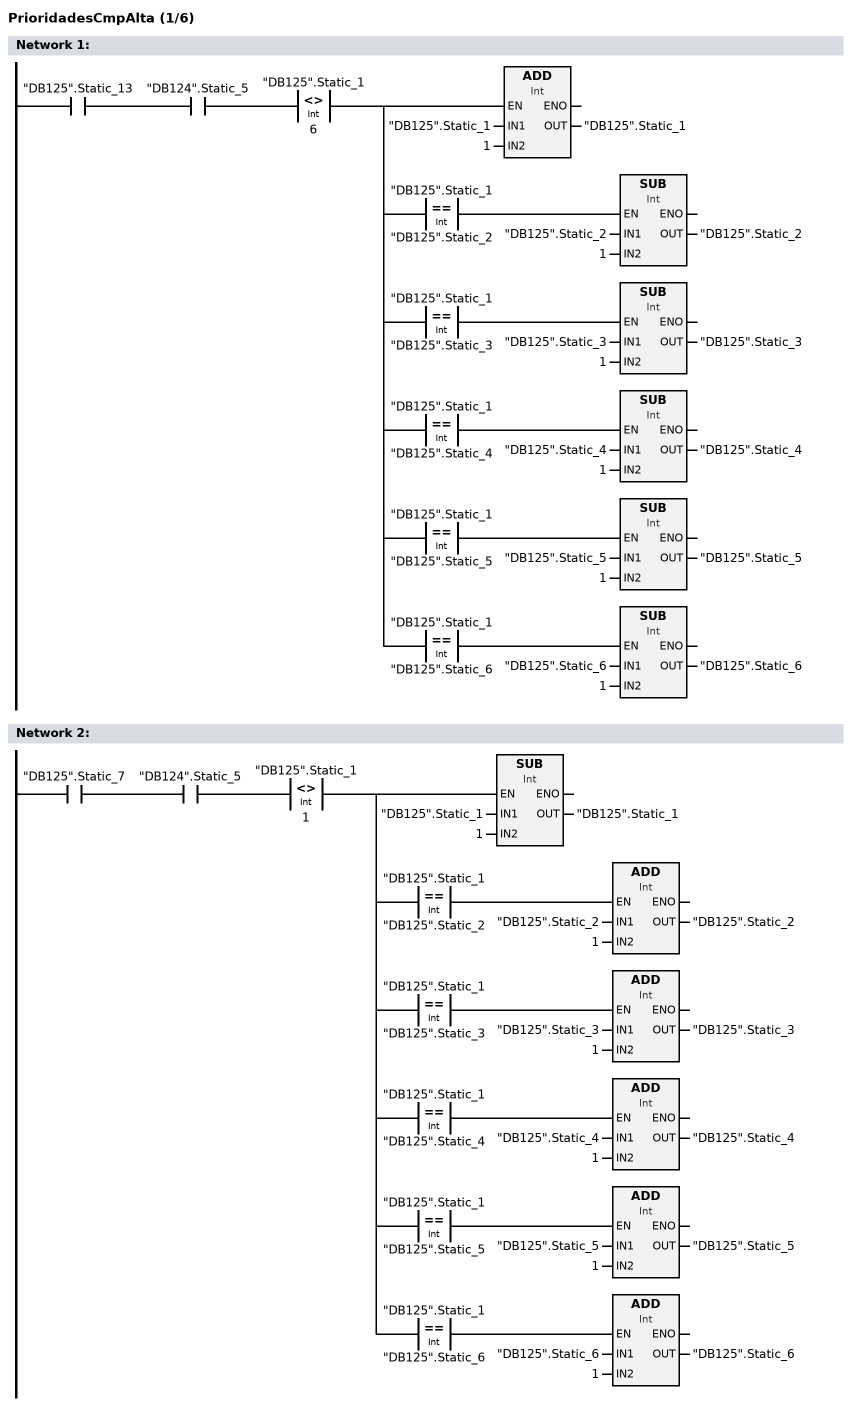
   #_w1 := "DB125".Static_13 AND "DB124".Static_5 AND ("DB125".Static_1 <> 6);
   IF #_w1 THEN "DB125".Static_1 := "DB125".Static_1 + 1; END_IF;
   IF #_w1 AND ("DB125".Static_1 = "DB125".Static_2) THEN "DB125".Static_2 := "DB125".Static_2 - 1; END_IF;
   IF #_w1 AND ("DB125".Static_1 = "DB125".Static_3) THEN "DB125".Static_3 := "DB125".Static_3 - 1; END_IF;
   IF #_w1 AND ("DB125".Static_1 = "DB125".Static_4) THEN "DB125".Static_4 := "DB125".Static_4 - 1; END_IF;
   IF #_w1 AND ("DB125".Static_1 = "DB125".Static_5) THEN "DB125".Static_5 := "DB125".Static_5 - 1; END_IF;
   IF #_w1 AND ("DB125".Static_1 = "DB125".Static_6) THEN "DB125".Static_6 := "DB125".Static_6 - 1; END_IF;
END_REGION

REGION Network 2
   #_w1 := "DB125".Static_7 AND "DB124".Static_5 AND ("DB125".Static_1 <> 1);
   IF #_w1 THEN "DB125".Static_1 := "DB125".Static_1 - 1; END_IF;
   IF #_w1 AND ("DB125".Static_1 = "DB125".Static_2) THEN "DB125".Static_2 := "DB125".Static_2 + 1; END_IF;
   IF #_w1 AND ("DB125".Static_1 = "DB125".Static_3) THEN "DB125".Static_3 := "DB125".Static_3 + 1; END_IF;
   IF #_w1 AND ("DB125".Static_1 = "DB125".Static_4) THEN "DB125".Static_4 := "DB125".Static_4 + 1; END_IF;
   IF #_w1 AND ("DB125".Static_1 = "DB125".Static_5) THEN "DB125".Static_5 := "DB125".Static_5 + 1; END_IF;
   IF #_w1 AND ("DB125".Static_1 = "DB125".Static_6) THEN "DB125".Static_6 := "DB125".Static_6 + 1; END_IF;
END_REGION

REGION Network 3
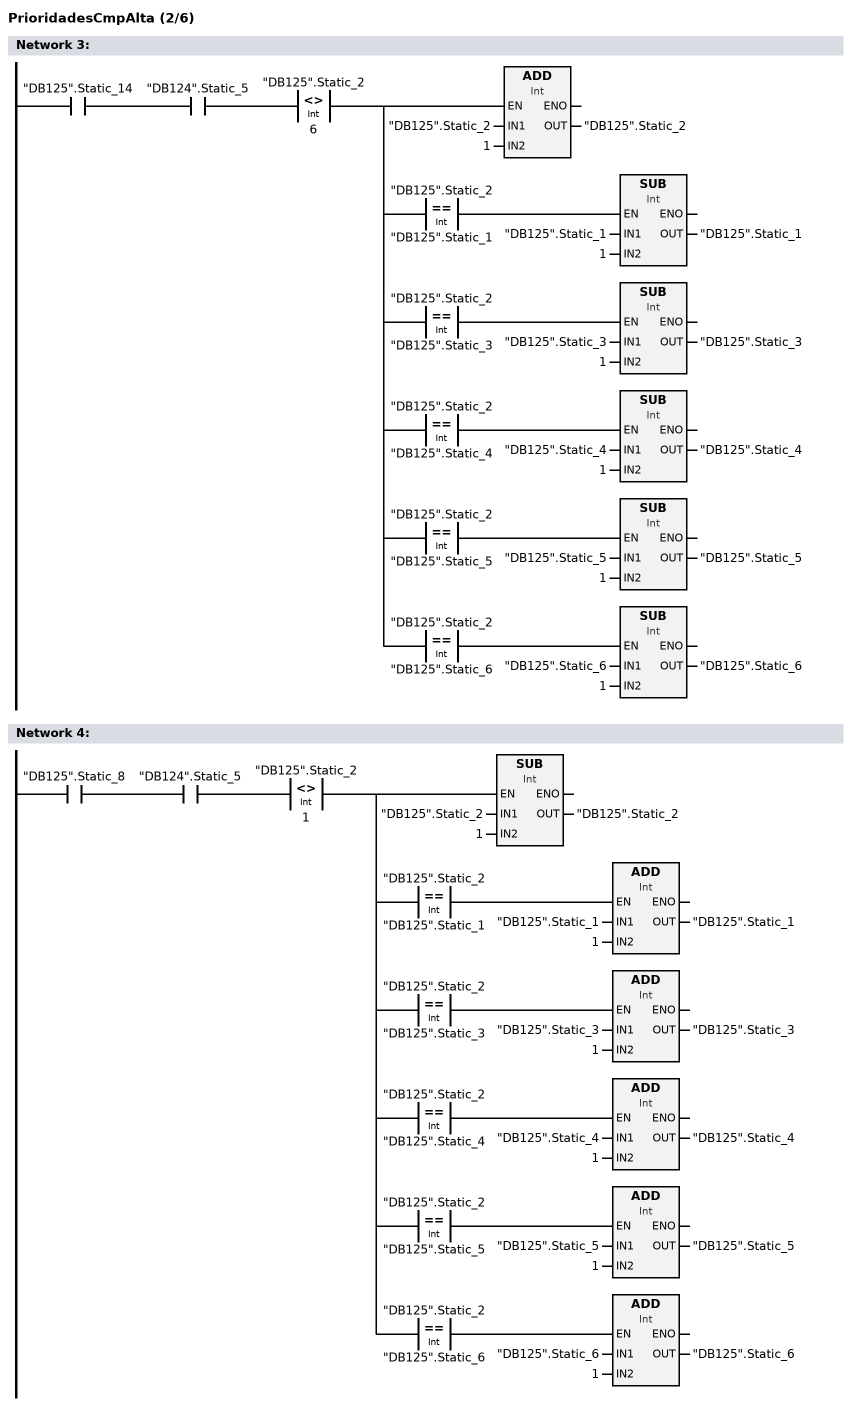
   #_w1 := "DB125".Static_14 AND "DB124".Static_5 AND ("DB125".Static_2 <> 6);
   IF #_w1 THEN "DB125".Static_2 := "DB125".Static_2 + 1; END_IF;
   IF #_w1 AND ("DB125".Static_2 = "DB125".Static_1) THEN "DB125".Static_1 := "DB125".Static_1 - 1; END_IF;
   IF #_w1 AND ("DB125".Static_2 = "DB125".Static_3) THEN "DB125".Static_3 := "DB125".Static_3 - 1; END_IF;
   IF #_w1 AND ("DB125".Static_2 = "DB125".Static_4) THEN "DB125".Static_4 := "DB125".Static_4 - 1; END_IF;
   IF #_w1 AND ("DB125".Static_2 = "DB125".Static_5) THEN "DB125".Static_5 := "DB125".Static_5 - 1; END_IF;
   IF #_w1 AND ("DB125".Static_2 = "DB125".Static_6) THEN "DB125".Static_6 := "DB125".Static_6 - 1; END_IF;
END_REGION

REGION Network 4
   #_w1 := "DB125".Static_8 AND "DB124".Static_5 AND ("DB125".Static_2 <> 1);
   IF #_w1 THEN "DB125".Static_2 := "DB125".Static_2 - 1; END_IF;
   IF #_w1 AND ("DB125".Static_2 = "DB125".Static_1) THEN "DB125".Static_1 := "DB125".Static_1 + 1; END_IF;
   IF #_w1 AND ("DB125".Static_2 = "DB125".Static_3) THEN "DB125".Static_3 := "DB125".Static_3 + 1; END_IF;
   IF #_w1 AND ("DB125".Static_2 = "DB125".Static_4) THEN "DB125".Static_4 := "DB125".Static_4 + 1; END_IF;
   IF #_w1 AND ("DB125".Static_2 = "DB125".Static_5) THEN "DB125".Static_5 := "DB125".Static_5 + 1; END_IF;
   IF #_w1 AND ("DB125".Static_2 = "DB125".Static_6) THEN "DB125".Static_6 := "DB125".Static_6 + 1; END_IF;
END_REGION

REGION Network 5
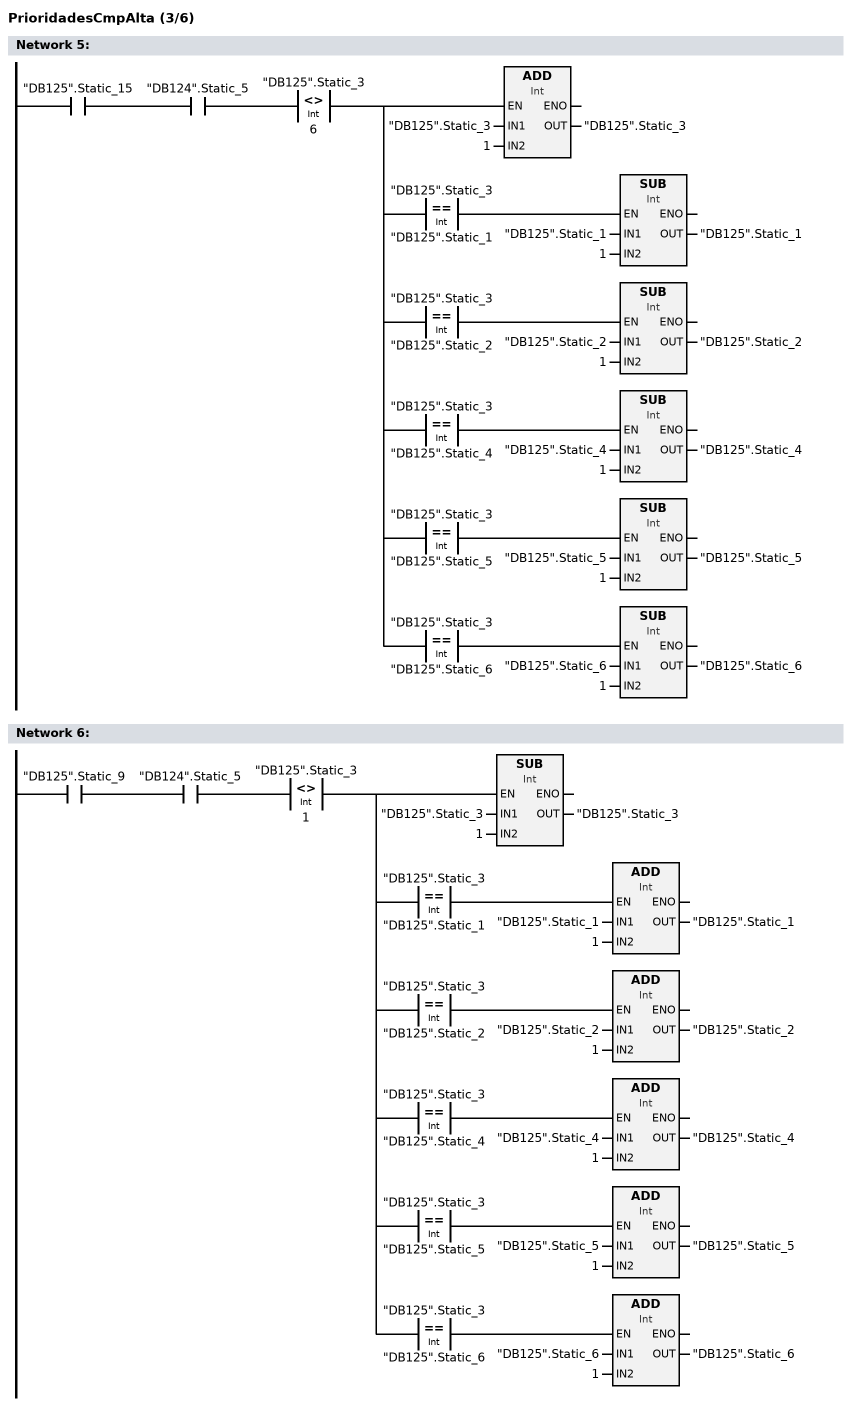
   #_w1 := "DB125".Static_15 AND "DB124".Static_5 AND ("DB125".Static_3 <> 6);
   IF #_w1 THEN "DB125".Static_3 := "DB125".Static_3 + 1; END_IF;
   IF #_w1 AND ("DB125".Static_3 = "DB125".Static_1) THEN "DB125".Static_1 := "DB125".Static_1 - 1; END_IF;
   IF #_w1 AND ("DB125".Static_3 = "DB125".Static_2) THEN "DB125".Static_2 := "DB125".Static_2 - 1; END_IF;
   IF #_w1 AND ("DB125".Static_3 = "DB125".Static_4) THEN "DB125".Static_4 := "DB125".Static_4 - 1; END_IF;
   IF #_w1 AND ("DB125".Static_3 = "DB125".Static_5) THEN "DB125".Static_5 := "DB125".Static_5 - 1; END_IF;
   IF #_w1 AND ("DB125".Static_3 = "DB125".Static_6) THEN "DB125".Static_6 := "DB125".Static_6 - 1; END_IF;
END_REGION

REGION Network 6
   #_w1 := "DB125".Static_9 AND "DB124".Static_5 AND ("DB125".Static_3 <> 1);
   IF #_w1 THEN "DB125".Static_3 := "DB125".Static_3 - 1; END_IF;
   IF #_w1 AND ("DB125".Static_3 = "DB125".Static_1) THEN "DB125".Static_1 := "DB125".Static_1 + 1; END_IF;
   IF #_w1 AND ("DB125".Static_3 = "DB125".Static_2) THEN "DB125".Static_2 := "DB125".Static_2 + 1; END_IF;
   IF #_w1 AND ("DB125".Static_3 = "DB125".Static_4) THEN "DB125".Static_4 := "DB125".Static_4 + 1; END_IF;
   IF #_w1 AND ("DB125".Static_3 = "DB125".Static_5) THEN "DB125".Static_5 := "DB125".Static_5 + 1; END_IF;
   IF #_w1 AND ("DB125".Static_3 = "DB125".Static_6) THEN "DB125".Static_6 := "DB125".Static_6 + 1; END_IF;
END_REGION

REGION Network 7
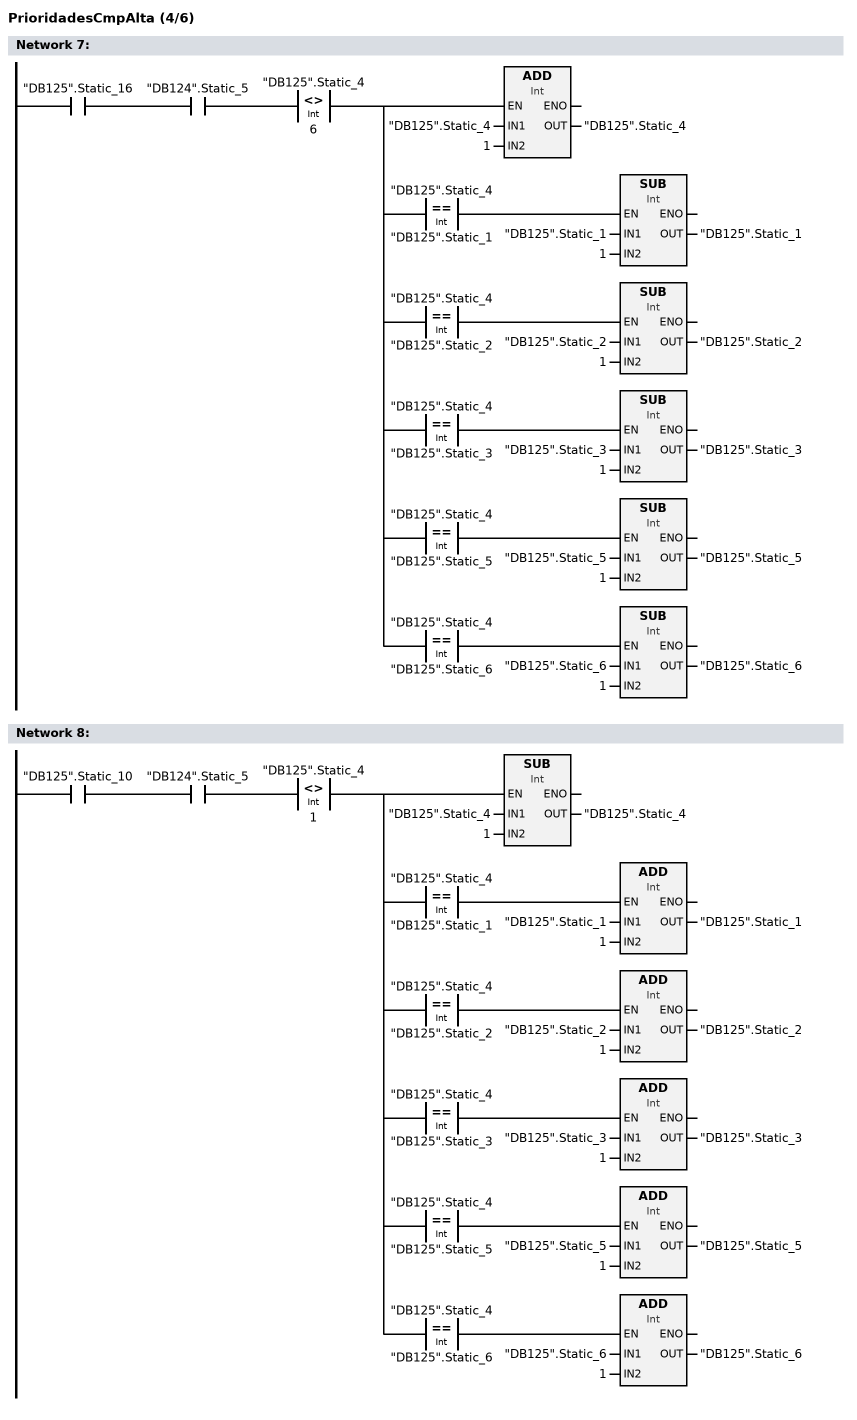
   #_w1 := "DB125".Static_16 AND "DB124".Static_5 AND ("DB125".Static_4 <> 6);
   IF #_w1 THEN "DB125".Static_4 := "DB125".Static_4 + 1; END_IF;
   IF #_w1 AND ("DB125".Static_4 = "DB125".Static_1) THEN "DB125".Static_1 := "DB125".Static_1 - 1; END_IF;
   IF #_w1 AND ("DB125".Static_4 = "DB125".Static_2) THEN "DB125".Static_2 := "DB125".Static_2 - 1; END_IF;
   IF #_w1 AND ("DB125".Static_4 = "DB125".Static_3) THEN "DB125".Static_3 := "DB125".Static_3 - 1; END_IF;
   IF #_w1 AND ("DB125".Static_4 = "DB125".Static_5) THEN "DB125".Static_5 := "DB125".Static_5 - 1; END_IF;
   IF #_w1 AND ("DB125".Static_4 = "DB125".Static_6) THEN "DB125".Static_6 := "DB125".Static_6 - 1; END_IF;
END_REGION

REGION Network 8
   #_w1 := "DB125".Static_10 AND "DB124".Static_5 AND ("DB125".Static_4 <> 1);
   IF #_w1 THEN "DB125".Static_4 := "DB125".Static_4 - 1; END_IF;
   IF #_w1 AND ("DB125".Static_4 = "DB125".Static_1) THEN "DB125".Static_1 := "DB125".Static_1 + 1; END_IF;
   IF #_w1 AND ("DB125".Static_4 = "DB125".Static_2) THEN "DB125".Static_2 := "DB125".Static_2 + 1; END_IF;
   IF #_w1 AND ("DB125".Static_4 = "DB125".Static_3) THEN "DB125".Static_3 := "DB125".Static_3 + 1; END_IF;
   IF #_w1 AND ("DB125".Static_4 = "DB125".Static_5) THEN "DB125".Static_5 := "DB125".Static_5 + 1; END_IF;
   IF #_w1 AND ("DB125".Static_4 = "DB125".Static_6) THEN "DB125".Static_6 := "DB125".Static_6 + 1; END_IF;
END_REGION

REGION Network 9
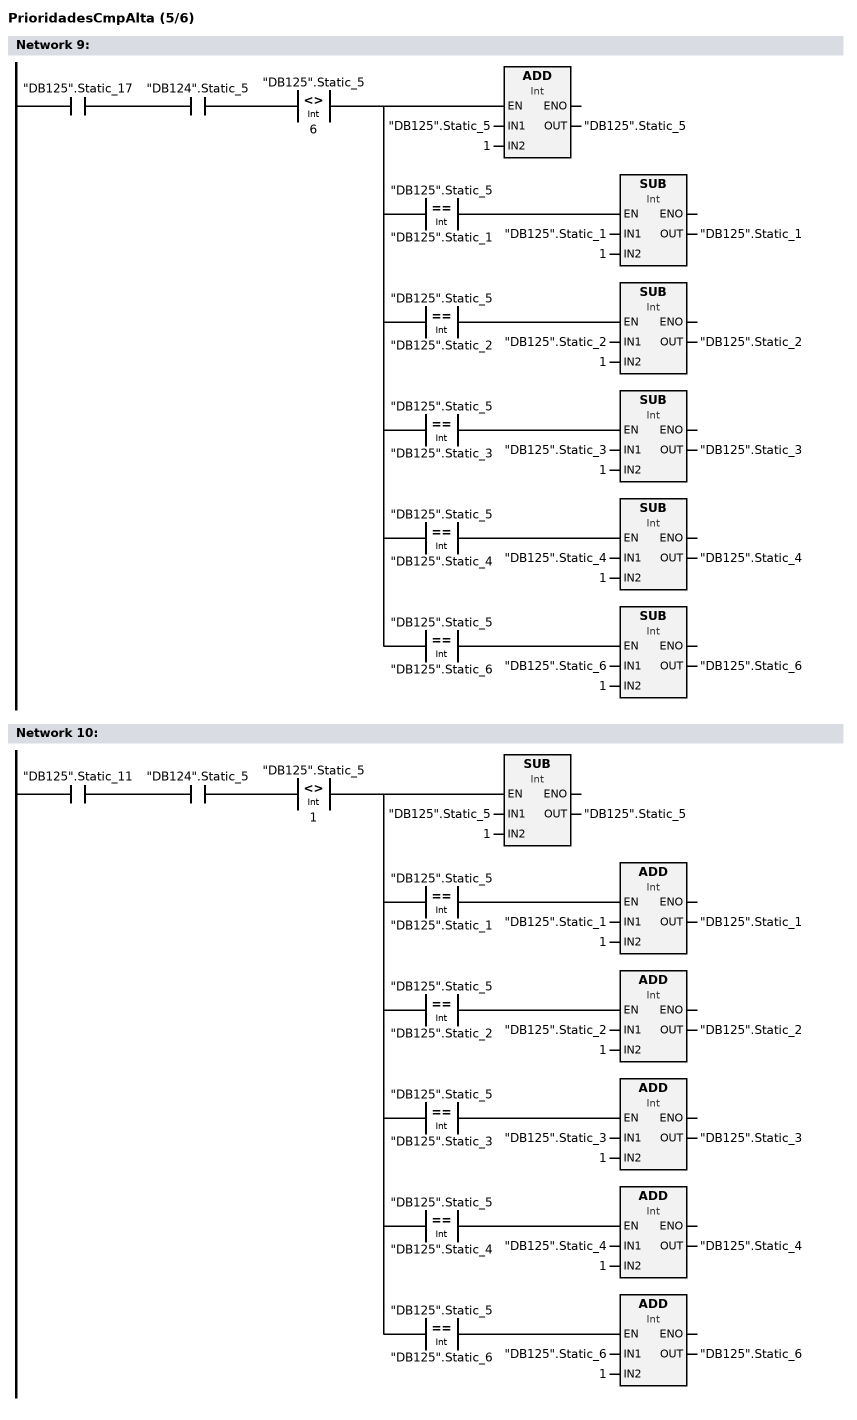
   #_w1 := "DB125".Static_17 AND "DB124".Static_5 AND ("DB125".Static_5 <> 6);
   IF #_w1 THEN "DB125".Static_5 := "DB125".Static_5 + 1; END_IF;
   IF #_w1 AND ("DB125".Static_5 = "DB125".Static_1) THEN "DB125".Static_1 := "DB125".Static_1 - 1; END_IF;
   IF #_w1 AND ("DB125".Static_5 = "DB125".Static_2) THEN "DB125".Static_2 := "DB125".Static_2 - 1; END_IF;
   IF #_w1 AND ("DB125".Static_5 = "DB125".Static_3) THEN "DB125".Static_3 := "DB125".Static_3 - 1; END_IF;
   IF #_w1 AND ("DB125".Static_5 = "DB125".Static_4) THEN "DB125".Static_4 := "DB125".Static_4 - 1; END_IF;
   IF #_w1 AND ("DB125".Static_5 = "DB125".Static_6) THEN "DB125".Static_6 := "DB125".Static_6 - 1; END_IF;
END_REGION

REGION Network 10
   #_w1 := "DB125".Static_11 AND "DB124".Static_5 AND ("DB125".Static_5 <> 1);
   IF #_w1 THEN "DB125".Static_5 := "DB125".Static_5 - 1; END_IF;
   IF #_w1 AND ("DB125".Static_5 = "DB125".Static_1) THEN "DB125".Static_1 := "DB125".Static_1 + 1; END_IF;
   IF #_w1 AND ("DB125".Static_5 = "DB125".Static_2) THEN "DB125".Static_2 := "DB125".Static_2 + 1; END_IF;
   IF #_w1 AND ("DB125".Static_5 = "DB125".Static_3) THEN "DB125".Static_3 := "DB125".Static_3 + 1; END_IF;
   IF #_w1 AND ("DB125".Static_5 = "DB125".Static_4) THEN "DB125".Static_4 := "DB125".Static_4 + 1; END_IF;
   IF #_w1 AND ("DB125".Static_5 = "DB125".Static_6) THEN "DB125".Static_6 := "DB125".Static_6 + 1; END_IF;
END_REGION

REGION Network 11
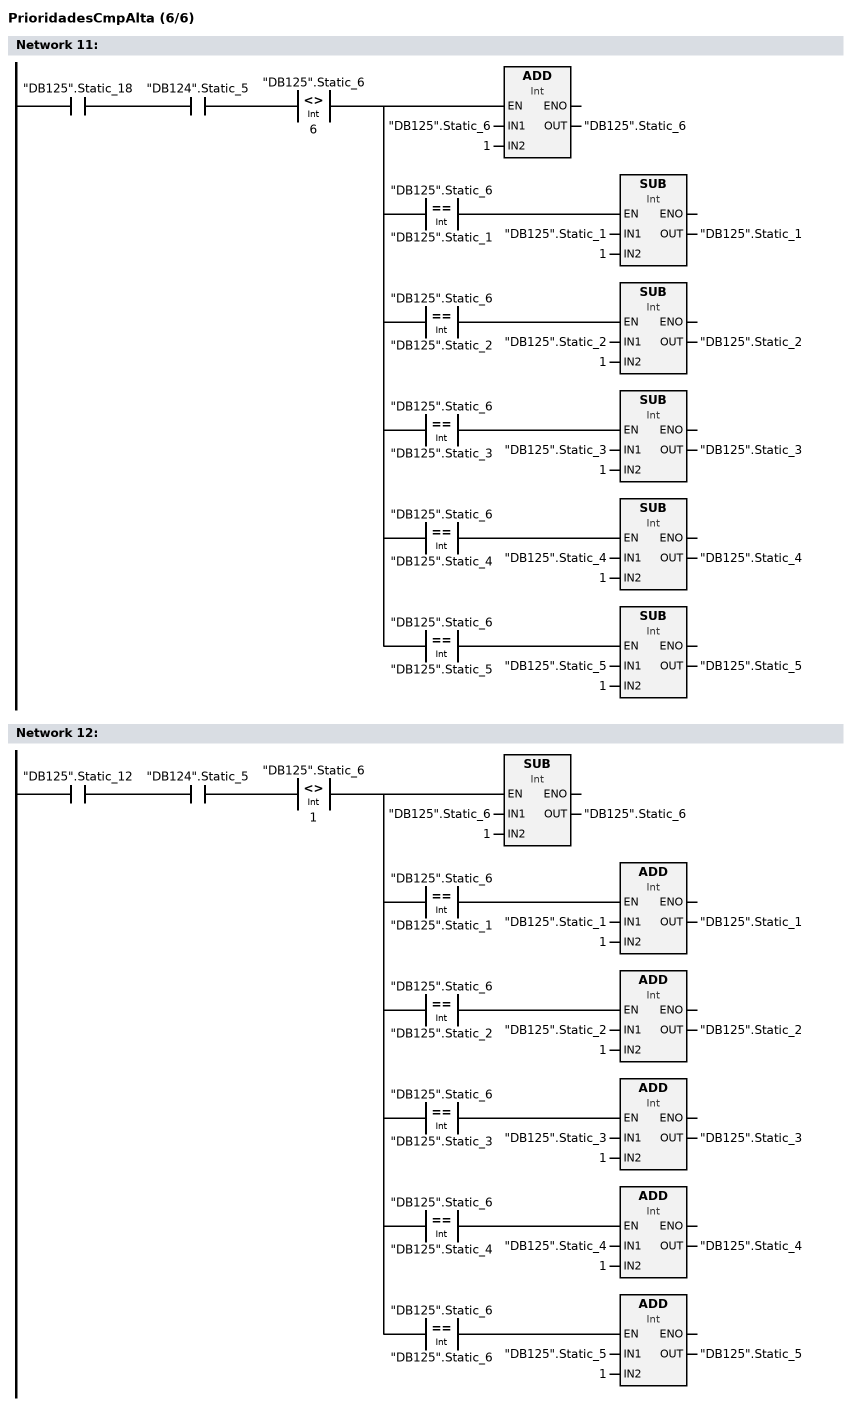
   #_w1 := "DB125".Static_18 AND "DB124".Static_5 AND ("DB125".Static_6 <> 6);
   IF #_w1 THEN "DB125".Static_6 := "DB125".Static_6 + 1; END_IF;
   IF #_w1 AND ("DB125".Static_6 = "DB125".Static_1) THEN "DB125".Static_1 := "DB125".Static_1 - 1; END_IF;
   IF #_w1 AND ("DB125".Static_6 = "DB125".Static_2) THEN "DB125".Static_2 := "DB125".Static_2 - 1; END_IF;
   IF #_w1 AND ("DB125".Static_6 = "DB125".Static_3) THEN "DB125".Static_3 := "DB125".Static_3 - 1; END_IF;
   IF #_w1 AND ("DB125".Static_6 = "DB125".Static_4) THEN "DB125".Static_4 := "DB125".Static_4 - 1; END_IF;
   IF #_w1 AND ("DB125".Static_6 = "DB125".Static_5) THEN "DB125".Static_5 := "DB125".Static_5 - 1; END_IF;
END_REGION

REGION Network 12
   #_w1 := "DB125".Static_12 AND "DB124".Static_5 AND ("DB125".Static_6 <> 1);
   IF #_w1 THEN "DB125".Static_6 := "DB125".Static_6 - 1; END_IF;
   IF #_w1 AND ("DB125".Static_6 = "DB125".Static_1) THEN "DB125".Static_1 := "DB125".Static_1 + 1; END_IF;
   IF #_w1 AND ("DB125".Static_6 = "DB125".Static_2) THEN "DB125".Static_2 := "DB125".Static_2 + 1; END_IF;
   IF #_w1 AND ("DB125".Static_6 = "DB125".Static_3) THEN "DB125".Static_3 := "DB125".Static_3 + 1; END_IF;
   IF #_w1 AND ("DB125".Static_6 = "DB125".Static_4) THEN "DB125".Static_4 := "DB125".Static_4 + 1; END_IF;
   IF #_w1 AND ("DB125".Static_6 = "DB125".Static_6) THEN "DB125".Static_5 := "DB125".Static_5 + 1; END_IF;
END_REGION
END_FUNCTION

FUNCTION "AccionamientosCmpAlta" : Void   // FC34, LAD
{ S7_Optimized_Access := 'FALSE' }
VERSION : 0.1
   VAR_TEMP   // added for the SCL form of the ladder/FBD networks
      _w1 : Bool;
      _s5time1 : S5Time;
   END_VAR
BEGIN

REGION Network 1
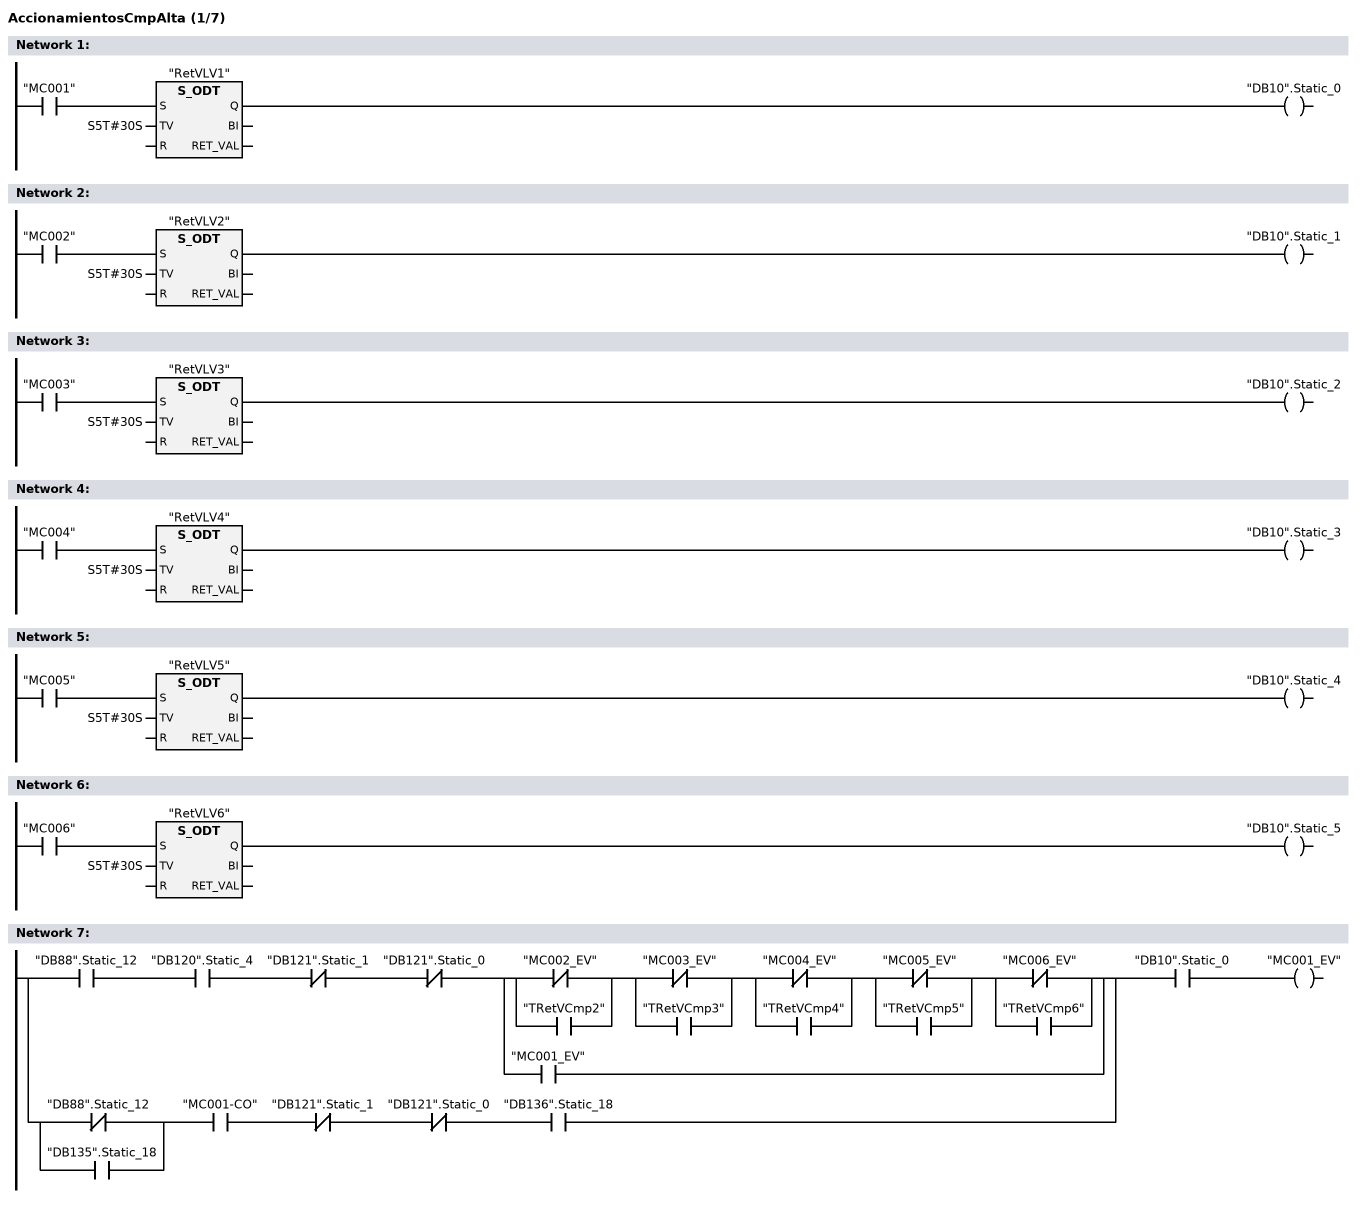
   RUNG wire#powerrail
      Contact( "MC001" )
      S_ODT(T_NO := "RetVLV1", TV := S5T#30S, R :=, BI =>, RET_VAL =>)
      Coil( "DB10".Static_0 )
   END_RUNG
   // the same network as SCL:
   #_s5time1 := S_ODT(T_NO := "RetVLV1", TV := S5T#30S, S := "MC001", Q => #_w1);
   "DB10".Static_0 := #_w1;
END_REGION

REGION Network 2
   RUNG wire#powerrail
      Contact( "MC002" )
      S_ODT(T_NO := "RetVLV2", TV := S5T#30S, R :=, BI =>, RET_VAL =>)
      Coil( "DB10".Static_1 )
   END_RUNG
   // the same network as SCL:
   #_s5time1 := S_ODT(T_NO := "RetVLV2", TV := S5T#30S, S := "MC002", Q => #_w1);
   "DB10".Static_1 := #_w1;
END_REGION

REGION Network 3
   RUNG wire#powerrail
      Contact( "MC003" )
      S_ODT(T_NO := "RetVLV3", TV := S5T#30S, R :=, BI =>, RET_VAL =>)
      Coil( "DB10".Static_2 )
   END_RUNG
   // the same network as SCL:
   #_s5time1 := S_ODT(T_NO := "RetVLV3", TV := S5T#30S, S := "MC003", Q => #_w1);
   "DB10".Static_2 := #_w1;
END_REGION

REGION Network 4
   RUNG wire#powerrail
      Contact( "MC004" )
      S_ODT(T_NO := "RetVLV4", TV := S5T#30S, R :=, BI =>, RET_VAL =>)
      Coil( "DB10".Static_3 )
   END_RUNG
   // the same network as SCL:
   #_s5time1 := S_ODT(T_NO := "RetVLV4", TV := S5T#30S, S := "MC004", Q => #_w1);
   "DB10".Static_3 := #_w1;
END_REGION

REGION Network 5
   RUNG wire#powerrail
      Contact( "MC005" )
      S_ODT(T_NO := "RetVLV5", TV := S5T#30S, R :=, BI =>, RET_VAL =>)
      Coil( "DB10".Static_4 )
   END_RUNG
   // the same network as SCL:
   #_s5time1 := S_ODT(T_NO := "RetVLV5", TV := S5T#30S, S := "MC005", Q => #_w1);
   "DB10".Static_4 := #_w1;
END_REGION

REGION Network 6
   RUNG wire#powerrail
      Contact( "MC006" )
      S_ODT(T_NO := "RetVLV6", TV := S5T#30S, R :=, BI =>, RET_VAL =>)
      Coil( "DB10".Static_5 )
   END_RUNG
   // the same network as SCL:
   #_s5time1 := S_ODT(T_NO := "RetVLV6", TV := S5T#30S, S := "MC006", Q => #_w1);
   "DB10".Static_5 := #_w1;
END_REGION

REGION Network 7
   "MC001_EV" := (("DB88".Static_12 AND "DB120".Static_4 AND NOT "DB121".Static_1 AND NOT "DB121".Static_0 AND (((NOT "MC002_EV" OR "TRetVCmp2") AND (NOT "MC003_EV" OR "TRetVCmp3") AND (NOT "MC004_EV" OR "TRetVCmp4") AND (NOT "MC005_EV" OR "TRetVCmp5") AND (NOT "MC006_EV" OR "TRetVCmp6")) OR "MC001_EV")) OR ((NOT "DB88".Static_12 OR "DB135".Static_18) AND "MC001-CO" AND NOT "DB121".Static_1 AND NOT "DB121".Static_0 AND "DB136".Static_18)) AND "DB10".Static_0;
END_REGION

REGION Network 8
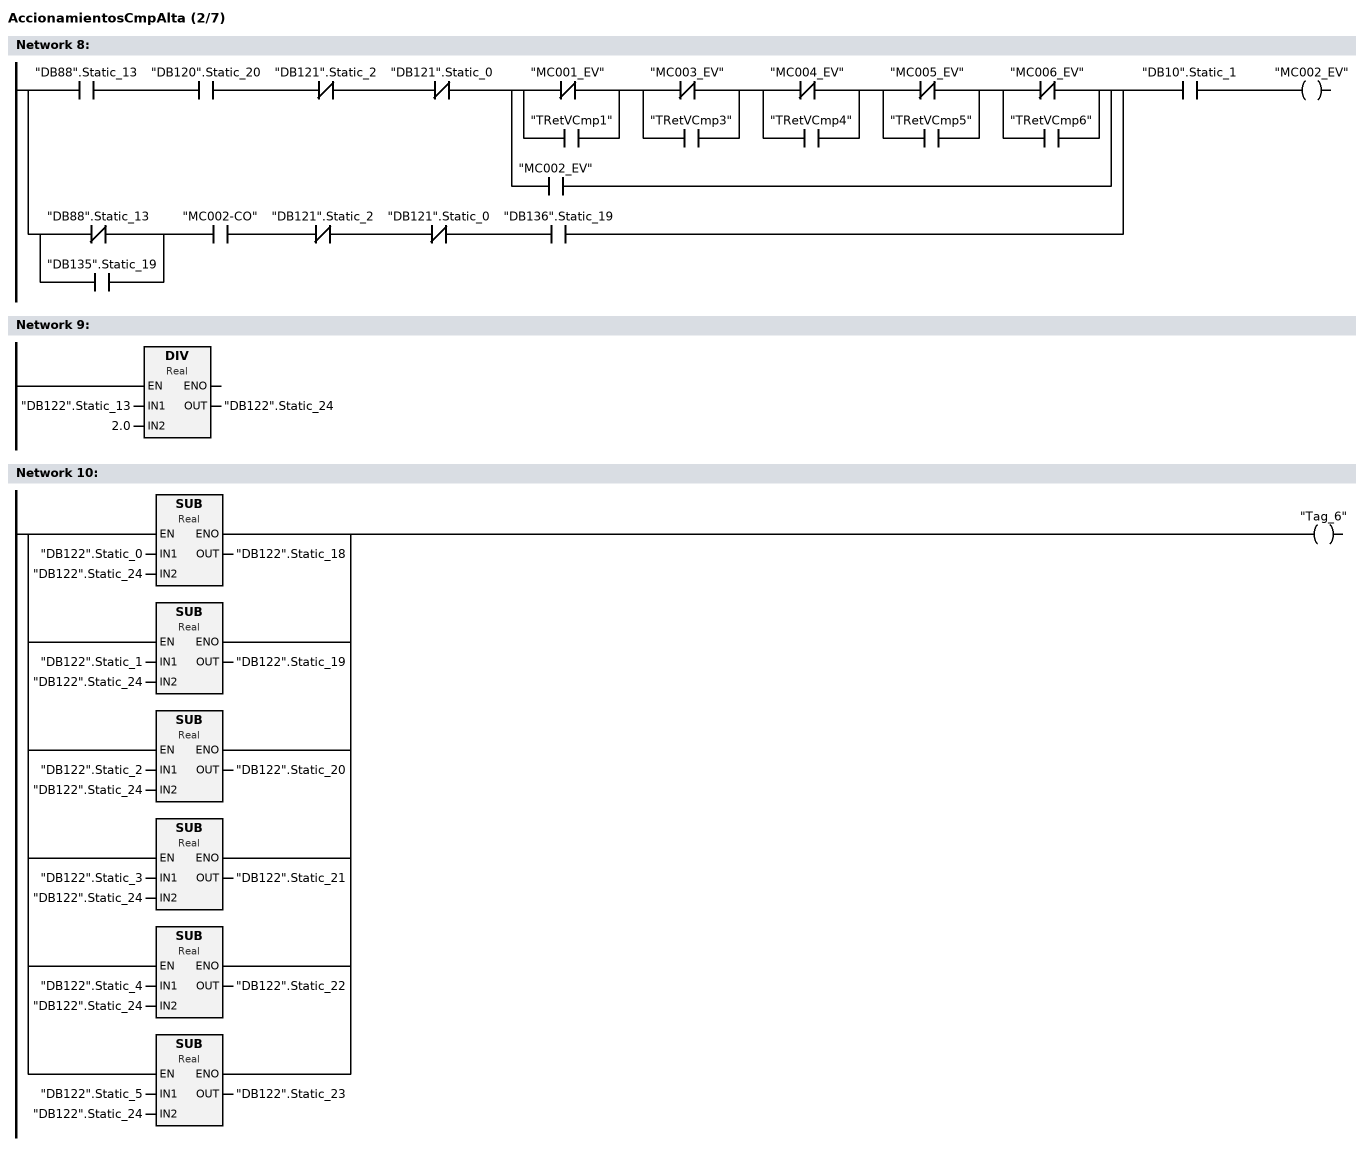
   "MC002_EV" := (("DB88".Static_13 AND "DB120".Static_20 AND NOT "DB121".Static_2 AND NOT "DB121".Static_0 AND (((NOT "MC001_EV" OR "TRetVCmp1") AND (NOT "MC003_EV" OR "TRetVCmp3") AND (NOT "MC004_EV" OR "TRetVCmp4") AND (NOT "MC005_EV" OR "TRetVCmp5") AND (NOT "MC006_EV" OR "TRetVCmp6")) OR "MC002_EV")) OR ((NOT "DB88".Static_13 OR "DB135".Static_19) AND "MC002-CO" AND NOT "DB121".Static_2 AND NOT "DB121".Static_0 AND "DB136".Static_19)) AND "DB10".Static_1;
END_REGION

REGION Network 9
   RUNG wire#powerrail
      { S7_Templates := "SrcType := Real"; S7_GenerateENO := "TRUE" } Div(in1 := "DB122".Static_13, in2 := 2.0, out => "DB122".Static_24)
   END_RUNG
   // the same network as SCL:
   "DB122".Static_24 := "DB122".Static_13 / 2.0;
END_REGION
